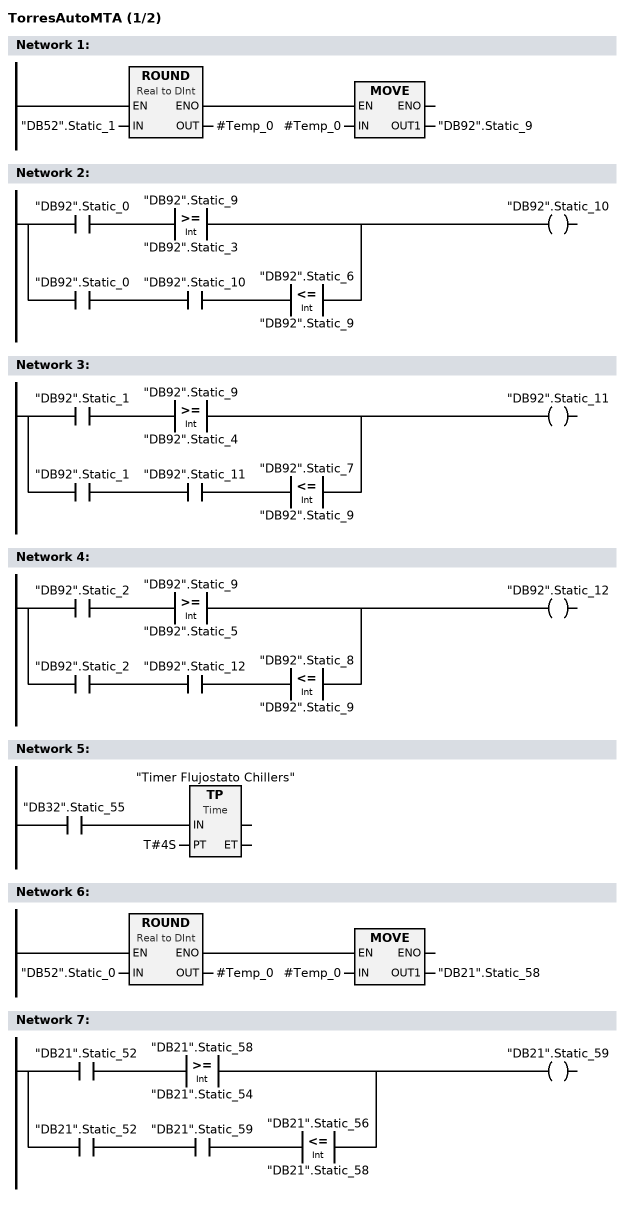
   RUNG wire#powerrail
      { S7_Templates := "[SrcType := Real, DestType := DInt]"; S7_GenerateENO := "TRUE" } Round(in := "DB52".Static_1, out => #Temp_0)
      { S7_GenerateENO := "TRUE" } Move(in := #Temp_0, out1 => "DB92".Static_9)
   END_RUNG
   // the same network as SCL:
   // ENO of a box is taken as its EN; it also drops when the box reports an error
   #Temp_0 := ROUND("DB52".Static_1);
   "DB92".Static_9 := #Temp_0;
END_REGION

REGION Network 2
   "DB92".Static_10 := ("DB92".Static_0 AND ("DB92".Static_9 >= "DB92".Static_3)) OR ("DB92".Static_0 AND "DB92".Static_10 AND ("DB92".Static_6 <= "DB92".Static_9));
END_REGION

REGION Network 3
   "DB92".Static_11 := ("DB92".Static_1 AND ("DB92".Static_9 >= "DB92".Static_4)) OR ("DB92".Static_1 AND "DB92".Static_11 AND ("DB92".Static_7 <= "DB92".Static_9));
END_REGION

REGION Network 4
   "DB92".Static_12 := ("DB92".Static_2 AND ("DB92".Static_9 >= "DB92".Static_5)) OR ("DB92".Static_2 AND "DB92".Static_12 AND ("DB92".Static_8 <= "DB92".Static_9));
END_REGION

REGION Network 5
   "Timer Flujostato Chillers".TP(pt := T#4S, in := "DB32".Static_55);
END_REGION

REGION Network 6
   RUNG wire#powerrail
      { S7_Templates := "[SrcType := Real, DestType := DInt]"; S7_GenerateENO := "TRUE" } Round(in := "DB52".Static_0, out => #Temp_0)
      { S7_GenerateENO := "TRUE" } Move(in := #Temp_0, out1 => "DB21".Static_58)
   END_RUNG
   // the same network as SCL:
   // ENO of a box is taken as its EN; it also drops when the box reports an error
   #Temp_0 := ROUND("DB52".Static_0);
   "DB21".Static_58 := #Temp_0;
END_REGION

REGION Network 7
   "DB21".Static_59 := ("DB21".Static_52 AND ("DB21".Static_58 >= "DB21".Static_54)) OR ("DB21".Static_52 AND "DB21".Static_59 AND ("DB21".Static_56 <= "DB21".Static_58));
END_REGION

REGION Network 8
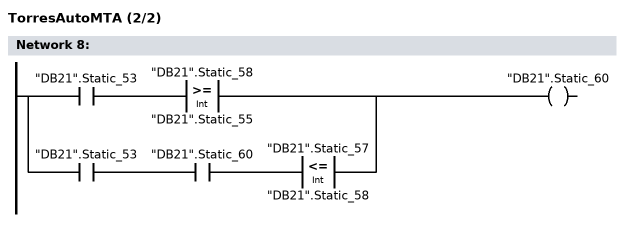
   "DB21".Static_60 := ("DB21".Static_53 AND ("DB21".Static_58 >= "DB21".Static_55)) OR ("DB21".Static_53 AND "DB21".Static_60 AND ("DB21".Static_57 <= "DB21".Static_58));
END_REGION
END_FUNCTION

(* ===== HMI "HMI_RT_3" =====
connection "Conexión2-PLC_1": ETHERNET, SIMATIC S7 300/400 MPI

HMI tags "AlarmasMTA"
   "AlarmasWord0" : Int, 1 s
   "AlarmasWord1" : Int, 1 s
   "AlarmasWord2" : Int, 1 s
   "AlarmasWord3" : Int, 1 s
   "AlarmasWord4" : Int, 1 s
   "AlarmasWord5" : Int, 1 s
   "AlarmasWord6" : Int, 1 s
   "AlarmasWord7" : Int, 1 s
   "AlarmasWord8" : Int, 1 s
   "Rec0" : Int, 1 s
   "Rec1" : Int, 1 s
   "Rec2" : Int, 1 s
   "Rec3" : Int, 1 s
   "Rec4" : Int, 1 s
   "Rec5" : Int, 1 s
   "Rec6" : Int, 1 s
   "Rec7" : Int, 1 s
   "Rec8" : Int, 1 s
   "AlarmasWord9" : Int, 1 s
   "AlarmasWord10" : Int, 1 s
   "AlarmasWord11" : Int, 1 s
   "AlarmasWord12" : Int, 1 s
   "AlarmasWord13" : Int, 1 s
   "AlarmasWord14" : Int, 1 s
   "Rec9" : Int, 1 s
   "Rec10" : Int, 1 s
   "Rec11" : Int, 1 s
   "Rec12" : Int, 1 s
   "Rec13" : Int, 1 s
   "Rec14" : Int, 1 s
   "AlarmasWord1(1)" : Int, 1 s
   "AlarmasWord15" : Int, 1 s
   "Rec15" : Int, 1 s
   "EncendidoPLC" : Bool, 1 s

HMI tags "AutoTorresChillers"
   "AutoV001" : Bool, 1 s
   "AutoV002" : Bool, 1 s
   "AutoV003" : Bool, 1 s
   "SP-ON-V001" : Int, 1 s
   "SP-ON-V002" : Int, 1 s
   "SP-ON-V003" : Int, 1 s
   "SP-OFF-V001" : Int, 1 s
   "SP-OFF-V002" : Int, 1 s
   "SP-OFF-V003" : Int, 1 s
   "TemperaturatorresCH" : Real, 1 s

HMI tags "CFG-Analog-MTA"
   "PresiónALTA" : Real, 1 s
   "PresiónBAJA" : Real, 1 s
   "TempCAV" : Real, 1 s
   "TempCH" : Real, 1 s
   "CFG-ALtaHH" : Real, 1 s
   "CFG-ALtaH" : Real, 1 s
   "CFG-ALtaL" : Real, 1 s
   "CFG-ALtaLL" : Real, 1 s
   "CFG-BajaHH" : Real, 1 s
   "CFG-BajaH" : Real, 1 s
   "CFG-BajaL" : Real, 1 s
   "CFG-BajaLL" : Real, 1 s

HMI tags "ChillersMTA"
   "HabMT007" : Bool, 1 s
   "HabMT008" : Bool, 1 s
   "HabMT009" : Bool, 1 s
   "HabMT010" : Bool, 1 s
   "DesMT007" : Bool, 1 s
   "DesMT008" : Bool, 1 s
   "DesMT009" : Bool, 1 s
   "DesMT010" : Bool, 1 s
   "MarchaMT007" : Bool, 1 s
   "MarchaMT008" : Bool, 1 s
   "MarchaMT009" : Bool, 1 s
   "MarchaMT010" : Bool, 1 s
   "ParadaMT007" : Bool, 1 s
   "ParadaMT008" : Bool, 1 s
   "ParadaMT009" : Bool, 1 s
   "ParadaMT010" : Bool, 1 s
   "Habilitación-CH-SOP-GR" : Bool, 1 s
   "Habilitación-CH-SOP-CH" : Bool, 1 s
   "Habilitación-CH-ENV-GR" : Bool, 1 s
   "Habilitación-CH-ENV-CH" : Bool, 1 s
   "Alarma1-CH-SOP-GR" : Bool, 1 s
   "Alarma2-CH-SOP-GR" : Bool, 1 s
   "RUN-CH-SOP-GR" : Bool, 1 s
   "MAX-CH-SOP-GR" : Bool, 1 s
   "AnimaciónMT007" : Byte, 1 s
   "AnimaciónMT008" : Byte, 1 s
   "AnimaciónMT009" : Byte, 1 s
   "AnimaciónMT010" : Byte, 1 s
   "AnimaciónMP010" : Byte, 1 s
   "AnimaciónMP011" : Byte, 1 s
   "AnimaciónMP012" : Byte, 1 s
   "AnimaciónMP013" : Byte, 1 s
   "HabMP010" : Bool, 1 s
   "HabMP011" : Bool, 1 s
   "HabMP012" : Bool, 1 s
   "HabMP013" : Bool, 1 s
   "HabMP018" : Bool, 1 s
   "HabMP019" : Bool, 1 s
   "DesMP010" : Bool, 1 s
   "DesMP011" : Bool, 1 s
   "DesMP012" : Bool, 1 s
   "DesMP013" : Bool, 1 s
   "DesMP018" : Bool, 1 s
   "DesMP019" : Bool, 1 s
   "MarchaMP010" : Bool, 1 s
   "MarchaMP011" : Bool, 1 s
   "MarchaMP012" : Bool, 1 s
   "MarchaMP013" : Bool, 1 s
   "MarchaMP018" : Bool, 1 s
   "MarchaMP019" : Bool, 1 s
   "ParadaMP010" : Bool, 1 s
   "ParadaMP011" : Bool, 1 s
   "ParadaMP012" : Bool, 1 s
   "ParadaMP013" : Bool, 1 s
   "ParadaMP018" : Bool, 1 s
   "ParadaMP019" : Bool, 1 s
   "AnimaciónMP018" : Byte, 1 s
   "AnimaciónMP019" : Byte, 1 s
   "DesV001" : Bool, 1 s
   "DesV002" : Bool, 1 s
   "HabV001" : Bool, 1 s
   "HabV002" : Bool, 1 s
   "MarchaV001" : Bool, 1 s
   "MarchaV002" : Bool, 1 s
   "ParadaV001" : Bool, 1 s
   "ParadaV002" : Bool, 1 s
   "AnimaciónV001" : Byte, 1 s
   "AnimaciónV002" : Byte, 1 s
   "VentiladoresMTA" : Bool, internal
   "MAX-CH-ENV-GR" : Bool, 1 s
   "RUN-CH-ENV-GR" : Bool, 1 s
   "Alarma2-CH-ENV-GR" : Bool, 1 s
   "Alarma1-CH-ENV-GR" : Bool, 1 s
   "SirenaM1" : Bool, 1 s
   "SirenaM2" : Bool, 1 s
   "SirenaM3" : Bool, 1 s
   "SirenaM4" : Bool, 1 s
   "AnimaciónV003" : Byte, 1 s
   "HabV003" : Bool, 1 s
   "DesV003" : Bool, 1 s
   "MarchaV003" : Bool, 1 s
   "ParadaV003" : Bool, 1 s
   "BombaTorreON" : Bool, 1 s
   "SirenaM5" : Bool, 1 s
   "SirenaChillers" : Bool, 1 s
   "SirenaM6" : Bool, 1 s
   "SirenaM7" : Bool, 1 s
   "SirenaM8" : Bool, 1 s
   "SirenaM9" : Bool, 1 s
   "SirenaM10" : Bool, 1 s
   "AlarmaNueva" : Bool, 1 s
   "AlarmaPresente" : Bool, 1 s
   "SinAlarmas" : Bool, 1 s
   "AlarmaAceite-CH-ENV-CH" : Bool, 1 s
   "AlarmaTemp-CH-ENV-CH" : Bool, 1 s
   "RUN-CH-ENV-CH" : Bool, 1 s
   "VerCh1MTA" : Bool, internal
   "VerCh2MTA" : Bool, internal
   "VerCh3MTA" : Bool, internal
   "VerCh4MTA" : Bool, internal
   "AlarmaPRUEBA" : DWord, 1 s
   "Presosato" : Bool, 1 s
   "CH-SOP-CH-CTC1ON" : Bool, 1 s
   "CH-SOP-CH-CTC2ON" : Bool, 1 s
   "CH-SOP-CH-TERM1" : Bool, 1 s
   "CH-SOP-CH-TERM2" : Bool, 1 s
   "CH-ENV-CH-ACT" : Bool, 1 s
   "CH-ENV-CH-TEMP" : Bool, 1 s
   "CH-ENV-CH-TERM" : Bool, 1 s
   "CH-ENV-CH-RUN" : Bool, 1 s
   "BombaTorreON2" : Bool, 1 s
   "HabV001(1)" : Bool, 1 s
   "HabV002(1)" : Bool, 1 s
   "HabV003(1)" : Bool, 1 s
   "HabV4" : Bool, 1 s
   "MarchaV001(1)" : Bool, 1 s
   "MarchaV002(1)" : Bool, 1 s
   "MarchaV003(1)" : Bool, 1 s
   "ParadaV001(1)" : Bool, 1 s
   "ParadaV002(1)" : Bool, 1 s
   "ParadaV003(1)" : Bool, 1 s
   "AnimaMenuV001" : Int, 1 s
   "AnimaMenuV002" : Int, 1 s
   "AnimaMenuV003" : Int, 1 s
   "DeshV001" : Bool, 1 s
   "DeshV002" : Bool, 1 s
   "DeshV003" : Bool, 1 s

discrete alarms
   125: '', class MTA, trigger "AlarmasWord4" bit 8
   126: '', class MTA, trigger "AlarmasWord3" bit 15
   127: '', class MTA, trigger "AlarmasWord4" bit 11
   128: '', class MTA, trigger "AlarmasWord4" bit 10
   129: '', class MTA, trigger "AlarmasWord4" bit 9
   130: '', class MTA, trigger "AlarmasWord3" bit 11
   131: '', class MTA, trigger "AlarmasWord3" bit 10
   132: '', class MTA, trigger "AlarmasWord3" bit 9
   133: '', class MTA, trigger "AlarmasWord3" bit 14
   134: '', class MTA, trigger "AlarmasWord3" bit 13
   135: '', class MTA, trigger "AlarmasWord3" bit 12
   136: '', class MTA, trigger "AlarmasWord4" bit 12
   137: '', class MTA, trigger "AlarmasWord4" bit 15
   138: '', class MTA, trigger "AlarmasWord4" bit 14
   139: '', class MTA, trigger "AlarmasWord4" bit 13
   140: '', class MTA, trigger "AlarmasWord3" bit 8
   141: '', class MTA, trigger "AlarmasWord1" bit 8
   144: '', class MTA, trigger "AlarmasWord1" bit 11
   145: '', class MTA, trigger "AlarmasWord1" bit 10
   146: '', class MTA, trigger "AlarmasWord1" bit 9
   153: '', class MTA, trigger "AlarmasWord1" bit 12
   154: '', class MTA, trigger "AlarmasWord2" bit 12
   155: '', class MTA, trigger "AlarmasWord2" bit 11
   156: '', class MTA, trigger "AlarmasWord2" bit 10
   157: '', class MTA, trigger "AlarmasWord2" bit 15
   158: '', class MTA, trigger "AlarmasWord2" bit 14
   159: '', class MTA, trigger "AlarmasWord2" bit 13
   160: '', class MTA, trigger "AlarmasWord1" bit 15
   161: '', class MTA, trigger "AlarmasWord1" bit 14
   162: '', class MTA, trigger "AlarmasWord1" bit 13
   163: '', class MTA, trigger "AlarmasWord2" bit 9
   164: '', class MTA, trigger "AlarmasWord2" bit 8
   165: '', class MTA, trigger "AlarmasWord5" bit 8
   166: '', class MTA, trigger "AlarmasWord5" bit 9
   167: '', class MTA, trigger "AlarmasWord5" bit 10
   168: '', class MTA, trigger "AlarmasWord5" bit 11
   169: '', class MTA, trigger "AlarmasWord5" bit 12
   170: '', class MTA, trigger "AlarmasWord5" bit 13
   171: '', class MTA, trigger "AlarmasWord5" bit 14
   172: '', class MTA, trigger "AlarmasWord5" bit 15
   13: '', class MTA, trigger "AlarmasWord6" bit 8
   14: '', class MTA, trigger "AlarmasWord6" bit 9
   50: '', class MTA, trigger "AlarmasWord6" bit 10
   53: '', class MTA, trigger "AlarmasWord6" bit 11
   87: '', class MTA, trigger "AlarmasWord6" bit 12
   88: '', class MTA, trigger "AlarmasWord6" bit 13
   89: '', class MTA, trigger "AlarmasWord6" bit 14
   90: '', class MTA, trigger "AlarmasWord6" bit 15
   69: '', class MTA, trigger "AlarmasWord7" bit 11
   68: '', class MTA, trigger "AlarmasWord7" bit 10
   67: '', class MTA, trigger "AlarmasWord7" bit 9
   66: '', class MTA, trigger "AlarmasWord7" bit 8
   70: '', class MTA, trigger "AlarmasWord7" bit 12
   71: '', class MTA, trigger "AlarmasWord7" bit 13
   72: '', class MTA, trigger "AlarmasWord7" bit 14
   73: '', class MTA, trigger "AlarmasWord7" bit 15
   74: '', class MTA, trigger "AlarmasWord8" bit 8
   75: '', class MTA, trigger "AlarmasWord8" bit 9
   76: '', class MTA, trigger "AlarmasWord8" bit 10
   77: '', class MTA, trigger "AlarmasWord8" bit 11
   78: '', class MTA, trigger "AlarmasWord8" bit 12
   79: '', class MTA, trigger "AlarmasWord8" bit 13
   80: '', class MTA, trigger "AlarmasWord8" bit 14
   81: '', class MTA, trigger "AlarmasWord8" bit 15
   82: '', class MTA, trigger "AlarmasWord9" bit 8
   83: '', class MTA, trigger "AlarmasWord9" bit 9
   91: '', class MTA, trigger "AlarmasWord9" bit 10
   92: '', class MTA, trigger "AlarmasWord9" bit 11
   93: '', class MTA, trigger "AlarmasWord9" bit 12
   94: '', class MTA, trigger "AlarmasWord9" bit 13
   96: '', class MTA, trigger "AlarmasWord9" bit 15
   97: '', class MTA, trigger "AlarmasWord10" bit 8
   98: '', class MTA, trigger "AlarmasWord10" bit 9
   99: '', class MTA, trigger "AlarmasWord10" bit 10
   100: '', class MTA, trigger "AlarmasWord10" bit 11
   101: '', class MTA, trigger "AlarmasWord10" bit 12
   102: '', class MTA, trigger "AlarmasWord10" bit 13
   121: '', class MTA, trigger "AlarmasWord10" bit 14
   104: '', class MTA, trigger "AlarmasWord10" bit 15
   105: '', class MTA, trigger "AlarmasWord11" bit 8
   106: '', class MTA, trigger "AlarmasWord11" bit 9
   107: '', class MTA, trigger "AlarmasWord11" bit 10
   108: '', class MTA, trigger "AlarmasWord11" bit 11
   109: '', class MTA, trigger "AlarmasWord11" bit 12
   110: '', class MTA, trigger "AlarmasWord11" bit 13
   111: '', class MTA, trigger "AlarmasWord11" bit 14
   112: '', class MTA, trigger "AlarmasWord11" bit 15
   113: '', class MTA, trigger "AlarmasWord12" bit 8
   114: '', class MTA, trigger "AlarmasWord12" bit 9
   115: '', class MTA, trigger "AlarmasWord12" bit 10
   116: '', class MTA, trigger "AlarmasWord12" bit 11
   117: '', class MTA, trigger "AlarmasWord12" bit 12
   118: '', class MTA, trigger "AlarmasWord12" bit 13
   119: '', class MTA, trigger "AlarmasWord12" bit 14
   120: '', class MTA, trigger "AlarmasWord12" bit 15
   122: '', class MTA, trigger "AlarmasWord13" bit 8
   1: '', class MTA, trigger "AlarmasWord13" bit 9
   2: '', class MTA, trigger "AlarmasWord13" bit 10
   3: '', class MTA, trigger "AlarmasWord13" bit 11
   4: '', class MTA, trigger "AlarmasWord13" bit 12
   5: '', class MTA, trigger "AlarmasWord13" bit 13
   6: '', class MTA, trigger "AlarmasWord13" bit 14
   7: '', class MTA, trigger "AlarmasWord13" bit 15
   8: '', class MTA, trigger "AlarmasWord14" bit 8
   9: '', class MTA, trigger "AlarmasWord14" bit 9
   10: '', class MTA, trigger "AlarmasWord14" bit 10
   11: '', class MTA, trigger "AlarmasWord14" bit 11
   12: '', class MTA, trigger "AlarmasWord14" bit 12
   15: '', class MTA, trigger "AlarmasWord14" bit 13
   16: '', class MTA, trigger "AlarmasWord14" bit 14
   17: '', class MTA, trigger "AlarmasWord14" bit 15
   95: '', class MTA, trigger "AlarmasWord9" bit 14
   149: '', class MTA, trigger "AlarmasWord0" bit 8
   142: '', class MTA, trigger "AlarmasWord0" bit 15
   143: '', class MTA, trigger "AlarmasWord0" bit 14
   152: '', class MTA, trigger "AlarmasWord0" bit 11
   147: '', class MTA, trigger "AlarmasWord0" bit 10
   148: '', class MTA, trigger "AlarmasWord0" bit 9
   150: '', class MTA, trigger "AlarmasWord0" bit 13
   151: '', class MTA, trigger "AlarmasWord0" bit 12
   21: '', class MTA, trigger "AlarmasWord15" bit 11
   22: '', class MTA, trigger "AlarmasWord15" bit 12
   19: '', class MTA, trigger "AlarmasWord15" bit 9
   20: '', class MTA, trigger "AlarmasWord15" bit 10
   23: '', class MTA, trigger "AlarmasWord15" bit 13
   24: '', class MTA, trigger "AlarmasWord15" bit 14
   25: '', class MTA, trigger "AlarmasWord15" bit 15
   18: '', class MTA, trigger "AlarmasWord15" bit 8

text list "EstadoMotor": 0 ''; 1 ''; 2 ''; 3 ''; 4 ''; 5 ''; 6 ''; 7 ''

graphic list "Motor2": 0 'Motor2Dorado'; 1 'Motor2Verde_1'; 2 'Motor2VerdeOscuro'; 3 'Motor2Azul'; 4 'Motor2Celeste'; 5 'Motor2Amarillo'; 6 'Motor2Gris_1'; 7 'Motor2Rojo'

graphic list "MotorTorre": 0 'torreFINAL4C2_1'; 1 'torreFINAL4C2v_2'; 2 'torreFINAL4C2v_2'; 3 'torreFINAL4C2b'; 4 'torreFINAL4C2b'; 5 'torreFINAL4C2a_2'; 6 'torreFINAL4C2_1'; 7 'torreFINAL4C2_1'

graphic list "Indicador": 0 'indDorado'; 1 'indVerde'; 2 'indVerde_1'; 3 'indAZUL'; 4 'indCeleste'; 5 'indAmarillo'; 6 'indGris'; 7 'indRojo'

graphic list "Secador2": 0 'BaseSullChicoDorado_2'; 1 'BaseSullChico_5'; 2 'BaseSullChico_5'; 3 'BaseSullChicoAzul_2'; 4 'BaseSullChicoAzul_2'; 5 'BaseSullChicoAmarillo_2'; 6 'BaseSullChicoGris_2'; 7 'BaseSullChicoRojo_2'

graphic list "Secador3": 0 'BaseSullChicoDorado_3'; 1 'BaseSullChico_6'; 2 'BaseSullChico_6'; 3 'BaseSullChicoAzul_3'; 4 'BaseSullChicoAzul_3'; 5 'BaseSullChicoAmarillo_3'; 6 'BaseSullChicoGris_3'; 7 'BaseSullChicoRojo_3'

graphic list "Secador1": 0 'BaseSullChicoDorado_1'; 1 'BaseSullChico_4'; 2 'BaseSullChico_4'; 3 'BaseSullChicoAzul_1'; 4 'BaseSullChicoAzul_1'; 5 'BaseSullChicoAmarillo_1'; 6 'BaseSullChicoGris_1'; 7 'BaseSullChicoRojo_1'

screen "MTA-Avisos" 800x480, template "Plantilla_2"
   AlarmView "Visor de avisos_1" at 5,53 size 790x367
   TextField "Campo de texto_5" at 327,10 size 54x27

screen "MTA-ChillersBombasEnvasado" 800x480, template "Plantilla_2"
   GraphicView "Visor de gráficos_3" at 648,158 size 48x71
   GraphicIOField "Plantilla_Campo ES gráfico_2" at 684,217 size 49x36
   SymbolicIOField "Campo ES simbólico_4" at 602,132 size 172x21
   TextField "Campo de texto_6" at 599,93 size 42x18
   GraphicView "Visor de gráficos_4" at 454,158 size 48x71
   GraphicIOField "Plantilla_Campo ES gráfico_1" at 490,217 size 49x36
   SymbolicIOField "Campo ES simbólico_1" at 408,132 size 172x21
   TextField "Campo de texto_7" at 405,93 size 42x18
   GraphicView "Visor de gráficos_6" at 64,158 size 48x71
   GraphicIOField "Plantilla_Campo ES gráfico_4" at 100,217 size 49x36
   SymbolicIOField "Campo ES simbólico_3" at 20,132 size 172x21
   TextField "Campo de texto_9" at 23,93 size 41x18
   TextField "Campo de texto_19" at 405,112 size 169x18
   GraphicView "Visor de gráficos_5" at 260,158 size 48x71
   GraphicIOField "Plantilla_Campo ES gráfico_3" at 296,217 size 49x36
   SymbolicIOField "Campo ES simbólico_2" at 214,132 size 172x21
   TextField "Campo de texto_8" at 211,93 size 41x18
   TextField "Campo de texto_18" at 598,112 size 150x18
   TextField "Campo de texto_16" at 215,113 size 150x18
   TextField "Campo de texto_17" at 21,113 size 146x18
   GraphicView "Plantilla_Visor de gráficos_2" at 752,6 size 35x35
   GraphicView "Plantilla_Visor de gráficos_1" at 752,6 size 35x35
   Button "Botón_1" at 740,1 size 57x44
   ScreenModuleView "ControlMotor-NoAUTO_1" at 609,271 size 163x76
   ScreenModuleView "ControlMotor-NoAUTO_2" at 413,271 size 163x76
   ScreenModuleView "ControlMotor-NoAUTO_3" at 219,271 size 163x76
   ScreenModuleView "ControlMotor-NoAUTO_4" at 22,271 size 163x76
   TextField "Campo de texto_5" at 256,10 size 261x27

screen "MTA-ChillersBombasSoplado" 800x480, template "Plantilla_2"
   TextField "Campo de texto_5" at 256,10 size 248x27
   GraphicView "Visor de gráficos_3" at 648,158 size 48x71
   GraphicIOField "Plantilla_Campo ES gráfico_8" at 684,217 size 49x36
   SymbolicIOField "Campo ES simbólico_4" at 602,132 size 172x21
   TextField "Campo de texto_6" at 599,93 size 42x18
   GraphicView "Visor de gráficos_4" at 454,158 size 48x71
   GraphicIOField "Plantilla_Campo ES gráfico_7" at 490,217 size 49x36
   SymbolicIOField "Campo ES simbólico_1" at 408,132 size 172x21
   TextField "Campo de texto_7" at 405,93 size 42x18
   GraphicView "Visor de gráficos_6" at 64,158 size 48x71
   GraphicIOField "Plantilla_Campo ES gráfico_5" at 100,217 size 49x36
   SymbolicIOField "Campo ES simbólico_3" at 20,132 size 172x21
   TextField "Campo de texto_9" at 23,93 size 41x18
   TextField "Campo de texto_19" at 407,113 size 140x18
   GraphicView "Visor de gráficos_5" at 260,158 size 48x71
   GraphicIOField "Plantilla_Campo ES gráfico_6" at 296,217 size 49x36
   SymbolicIOField "Campo ES simbólico_2" at 214,132 size 172x21
   TextField "Campo de texto_8" at 211,93 size 41x18
   TextField "Campo de texto_18" at 599,113 size 104x18
   TextField "Campo de texto_16" at 212,113 size 142x18
   TextField "Campo de texto_17" at 21,113 size 138x18
   GraphicView "Plantilla_Visor de gráficos_2" at 752,6 size 35x35
   GraphicView "Plantilla_Visor de gráficos_1" at 752,6 size 35x35
   Button "Botón_1" at 740,1 size 57x44
   ScreenModuleView "ControlMotor-NoAUTO_1" at 609,271 size 163x76
   ScreenModuleView "ControlMotor-NoAUTO_3" at 219,271 size 163x76
   ScreenModuleView "ControlMotor-NoAUTO_2" at 417,271 size 163x76
   ScreenModuleView "ControlMotor-NoAUTO_4" at 27,271 size 163x76

screen "MTA-ChillersConfiguraciónSirena" 800x480, template "Plantilla_2"
   Switch "Interruptor_1" at 119,81 size 36x32
   Switch "Interruptor_2" at 119,118 size 36x32
   Switch "Interruptor_3" at 119,155 size 36x32
   Switch "Interruptor_4" at 119,192 size 36x32
   Switch "Interruptor_5" at 119,229 size 36x32
   TextField "Campo de texto_1" at 163,233 size 365x22
   TextField "Campo de texto_2" at 163,196 size 424x22
   TextField "Campo de texto_3" at 163,160 size 353x22
   TextField "Campo de texto_4" at 163,122 size 411x22
   TextField "Campo de texto_5" at 163,86 size 340x22
   TextField "Campo de texto_6" at 51,53 size 277x22
   TextField "Campo de texto_7" at 214,8 size 319x29
   Switch "Interruptor_6" at 119,266 size 36x32
   TextField "Campo de texto_8" at 163,271 size 231x22
   Switch "Interruptor_7" at 119,303 size 36x32
   TextField "Campo de texto_9" at 163,307 size 244x22
   Switch "Interruptor_8" at 119,341 size 36x32
   TextField "Campo de texto_10" at 163,346 size 150x22
   GraphicView "Plantilla_Visor de gráficos_2" at 752,6 size 35x35
   GraphicView "Plantilla_Visor de gráficos_1" at 752,6 size 35x35
   Button "Botón_1" at 740,1 size 57x44
   Switch "Interruptor_9" at 119,378 size 36x32
   TextField "Campo de texto_11" at 163,383 size 194x22

screen "MTA-Chillers-Envasado" 800x480, template "Plantilla_2"
   GraphicView "Visor de gráficos_2" at 24,127 size 192x232
   GraphicView "Visor de gráficos_1" at 432,129 size 144x104
   Switch "Interruptor_1" at 243,127 size 91x31
   TextField "Campo de texto_5" at 309,10 size 182x27
   TextField "Campo de texto_10" at 19,78 size 169x22
   TextField "Campo de texto_6" at 411,78 size 158x22
   TextField "Campo de texto_1" at 263,203 size 40x18
   TextField "Campo de texto_3" at 263,182 size 108x18
   TextField "Campo de texto_4" at 263,223 size 101x18
   Switch "Interruptor_2" at 595,127 size 91x31
   GraphicView "Plantilla_Visor de gráficos_2" at 752,6 size 35x35
   GraphicView "Plantilla_Visor de gráficos_1" at 752,6 size 35x35
   Button "Botón_1" at 740,1 size 57x44
   TextField "Campo de texto_24" at 613,183 size 79x18
   TextField "Campo de texto_25" at 613,166 size 108x18
   TextField "Campo de texto_26" at 613,201 size 115x18
   TextField "Campo de texto_27" at 613,220 size 125x18

screen "MTA-Chillers-General" 800x480, template "Plantilla_2"
   GraphicView "Visor de gráficos_7" at 488,183 size 48x71
   GraphicView "Visor de gráficos_8" at 536,183 size 48x71
   GraphicView "Visor de gráficos_1" at 392,183 size 48x71
   GraphicView "Visor de gráficos_9" at 440,183 size 48x71
   GraphicView "Visor de gráficos_17" at 383,130 size 87x77
   GraphicView "Visor de gráficos_18" at 479,130 size 87x77
   GraphicView "Visor de gráficos_14" at 384,48 size 141x131
   GraphicView "Visor de gráficos_3" at 750,189 size 48x212
   GraphicView "Visor de gráficos_4" at 630,161 size 96x96
   GraphicView "Visor de gráficos_5" at 264,183 size 48x71
   GraphicView "Visor de gráficos_6" at 312,183 size 48x71
   GraphicView "Visor de gráficos_10" at 168,183 size 48x71
   GraphicView "Visor de gráficos_11" at 216,183 size 48x71
   GraphicView "Visor de gráficos_2" at 12,132 size 128x144
   GraphicView "Visor de gráficos_12" at 45,333 size 88x77
   GraphicView "Visor de gráficos_15" at 159,130 size 87x77
   GraphicView "Visor de gráficos_16" at 255,130 size 87x77
   GraphicView "Visor de gráficos_13" at 162,48 size 141x131
   GraphicIOField "Plantilla_Campo ES gráfico_2" at 304,240 size 41x36
   GraphicIOField "Plantilla_Campo ES gráfico_1" at 352,240 size 41x36
   GraphicIOField "Plantilla_Campo ES gráfico_3" at 528,240 size 41x36
   GraphicIOField "Plantilla_Campo ES gráfico_4" at 576,240 size 41x36
   GraphicIOField "Plantilla_Campo ES gráfico_5" at 432,240 size 41x36
   GraphicIOField "Plantilla_Campo ES gráfico_6" at 480,240 size 41x36
   GraphicIOField "Plantilla_Campo ES gráfico_7" at 208,240 size 41x36
   GraphicIOField "Plantilla_Campo ES gráfico_8" at 256,240 size 41x36
   TextField "Campo de texto_1" at 631,124 size 86x32
   TextField "Campo de texto_2" at 668,364 size 86x32
   TextField "Campo de texto_3" at 142,373 size 90x32
   TextField "Campo de texto_4" at 28,94 size 90x32
   TextField "Campo de texto_5" at 334,8 size 72x29
   TextField "Campo de texto_6" at 474,309 size 131x25
   TextField "Campo de texto_7" at 242,309 size 139x25
   TextField "Campo de texto_9" at 520,70 size 51x52
   TextField "Campo de texto_8" at 214,277 size 41x19
   TextField "Campo de texto_11" at 262,277 size 41x19
   TextField "Campo de texto_12" at 310,277 size 49x19
   TextField "Campo de texto_13" at 366,277 size 42x19
   TextField "Campo de texto_14" at 438,277 size 41x19
   TextField "Campo de texto_15" at 486,277 size 41x19
   TextField "Campo de texto_16" at 534,277 size 42x19
   TextField "Campo de texto_17" at 590,277 size 42x19
   TextField "Campo de texto_10" at 294,69 size 58x52
   Button "Botón_3" at 629,155 size 170x254
   Button "Botón_2" at 419,227 size 215x78
   Button "Botón_4" at 0,122 size 194x294
   Button "Botón_5" at 203,226 size 208x79
   GraphicView "Plantilla_Visor de gráficos_2" at 752,6 size 35x35
   GraphicView "Plantilla_Visor de gráficos_1" at 752,6 size 35x35
   Button "Botón_1" at 740,1 size 57x44

screen "MTA-Chillers-Soplado" 800x480, template "Plantilla_2"
   GraphicView "Visor de gráficos_2" at 24,127 size 192x232
   GraphicView "Visor de gráficos_1" at 424,129 size 160x168
   Switch "Interruptor_1" at 243,127 size 91x31
   TextField "Campo de texto_1" at 263,203 size 40x18
   TextField "Campo de texto_3" at 263,182 size 108x18
   TextField "Campo de texto_4" at 263,223 size 101x18
   TextField "Campo de texto_5" at 311,10 size 169x27
   TextField "Campo de texto_10" at 19,78 size 156x22
   TextField "Campo de texto_6" at 411,78 size 145x22
   Switch "Interruptor_2" at 627,127 size 91x31
   GraphicView "Plantilla_Visor de gráficos_2" at 752,6 size 35x35
   GraphicView "Plantilla_Visor de gráficos_1" at 752,6 size 35x35
   Button "Botón_1" at 740,1 size 57x44
   TextField "Campo de texto_28" at 607,198 size 120x18
   TextField "Campo de texto_29" at 607,177 size 120x18
   TextField "Campo de texto_30" at 631,220 size 96x18
   TextField "Campo de texto_31" at 631,241 size 96x18

screen "MTA-TorreEnfriamientoBMB" 800x480, template "Plantilla_2"
   GraphicView "Visor de gráficos_1" at 167,153 size 98x119
   GraphicView "Visor de gráficos_4" at 260,143 size 138x153
   GraphicView "Visor de gráficos_17" at 16,128 size 178x201
   GraphicView "Visor de gráficos_2" at 167,153 size 98x119
   GraphicView "Visor de gráficos_3" at 260,143 size 138x153
   GraphicView "Visor de gráficos_5" at 16,128 size 178x201
   GraphicView "Visor de gráficos_6" at 167,153 size 98x119
   GraphicView "Visor de gráficos_15" at 260,143 size 138x153
   GraphicView "Visor de gráficos_16" at 16,128 size 178x201
   TextField "Campo de texto_1" at 361,84 size 57x23
   TextField "Campo de texto_2" at 229,95 size 47x20
   TextField "Campo de texto_12" at 101,76 size 57x23
   TextField "Campo de texto_13" at 273,197 size 55x29
   TextField "Campo de texto_14" at 38,202 size 50x34
   GraphicIOField "Campo ES gráfico_1" at 76,122 size 56x29
   GraphicIOField "Campo ES gráfico_2" at 199,147 size 33x21
   GraphicIOField "Campo ES gráfico_3" at 306,137 size 45x24
   GraphicView "Visor de gráficos_19" at 0,384 size 800x15
   GraphicView "Plantilla_Visor de gráficos_2" at 752,6 size 35x35
   GraphicView "Plantilla_Visor de gráficos_1" at 752,6 size 35x35
   Button "Botón_1" at 740,1 size 57x44
   Button "Botón_2" at 200,320 size 152x38
   TextField "Campo de texto_10" at 41,374 size 98x32
   TextField "Campo de texto_5" at 238,8 size 293x29
   GraphicView "Visor de gráficos_9" at 30,56 size 63x62
   GraphicView "Visor de gráficos_10" at 30,56 size 63x62
   GraphicView "Visor de gráficos_11" at 177,82 size 47x46
   GraphicView "Visor de gráficos_12" at 177,82 size 47x46
   GraphicView "Visor de gráficos_13" at 292,66 size 63x62
   GraphicView "Visor de gráficos_14" at 292,66 size 63x62
   IOField "Campo ES_1" at 241,360 size 80x23
   GraphicView "Visor de gráficos_8" at 459,277 size 48x71
   GraphicIOField "Plantilla_Campo ES gráfico_1" at 497,336 size 49x36
   SymbolicIOField "Campo ES simbólico_1" at 581,259 size 172x20
   TextField "Campo de texto_7" at 495,293 size 41x18
   TextField "Campo de texto_17" at 455,241 size 129x27
   ScreenModuleView "ControlMotor-NoAUTO_4" at 565,285 size 203x76
   ScreenModuleView "ControlMotor-NoAUTO_1" at 564,115 size 203x76
   SymbolicIOField "Campo ES simbólico_4" at 575,89 size 172x20
   TextField "Campo de texto_6" at 494,129 size 41x18
   TextField "Campo de texto_16" at 454,77 size 151x27
   GraphicView "Visor de gráficos_7" at 458,113 size 48x71
   GraphicIOField "Plantilla_Campo ES gráfico_2" at 496,172 size 49x36

screen "MTA-TorreEnfriamientoVENT" 800x480, template "Plantilla_2"
   GraphicView "Visor de gráficos_1" at 167,153 size 98x119
   GraphicView "Visor de gráficos_4" at 260,143 size 138x153
   GraphicView "Visor de gráficos_17" at 16,128 size 178x201
   GraphicView "Visor de gráficos_2" at 167,153 size 98x119
   GraphicView "Visor de gráficos_3" at 260,143 size 138x153
   GraphicView "Visor de gráficos_5" at 16,128 size 178x201
   GraphicView "Visor de gráficos_6" at 167,153 size 98x119
   GraphicView "Visor de gráficos_15" at 260,143 size 138x153
   GraphicView "Visor de gráficos_16" at 16,128 size 178x201
   SymbolicIOField "Campo ES simbólico_2" at 548,59 size 188x19
   SymbolicIOField "Campo ES simbólico_3" at 549,181 size 188x19
   SymbolicIOField "Campo ES simbólico_7" at 549,301 size 188x19
   TextField "Campo de texto_1" at 361,84 size 57x23
   TextField "Campo de texto_2" at 229,95 size 47x20
   TextField "Campo de texto_13" at 273,197 size 55x29
   TextField "Campo de texto_14" at 38,202 size 50x34
   ScreenModuleView "Faceplate_4_1" at 447,84 size 245x68
   TextField "Campo de texto_4" at 439,176 size 104x27
   TextField "Campo de texto_3" at 439,54 size 104x27
   TextField "Campo de texto_23" at 440,298 size 104x27
   ScreenModuleView "Faceplate_4_2" at 447,204 size 245x68
   ScreenModuleView "Faceplate_4_3" at 447,326 size 245x68
   TextField "Campo de texto_12" at 101,76 size 57x23
   GraphicIOField "Campo ES gráfico_1" at 76,122 size 56x29
   GraphicIOField "Campo ES gráfico_2" at 199,147 size 33x21
   GraphicIOField "Campo ES gráfico_3" at 306,137 size 45x24
   Switch "Interruptor_1" at 744,62 size 32x29
   Switch "Interruptor_2" at 744,184 size 32x29
   Switch "Interruptor_3" at 744,304 size 32x29
   GraphicView "Visor de gráficos_19" at 0,384 size 800x15
   TextField "Campo de texto_5" at 238,8 size 293x29
   GraphicView "Visor de gráficos_9" at 30,56 size 63x62
   GraphicView "Visor de gráficos_10" at 30,56 size 63x62
   GraphicView "Visor de gráficos_11" at 177,82 size 47x46
   GraphicView "Visor de gráficos_12" at 177,82 size 47x46
   GraphicView "Visor de gráficos_13" at 292,66 size 63x62
   GraphicView "Visor de gráficos_14" at 292,66 size 63x62
   GraphicView "Plantilla_Visor de gráficos_2" at 752,6 size 35x35
   GraphicView "Plantilla_Visor de gráficos_1" at 752,6 size 35x35
   Button "Botón_1" at 740,1 size 57x44
   TextField "Campo de texto_10" at 41,374 size 98x32
   Button "Botón_2" at 200,320 size 152x38
   IOField "Campo ES_1" at 241,360 size 80x23
   GraphicIOField "Campo ES gráfico_4" at 429,160 size 362x6
   GraphicIOField "Campo ES gráfico_5" at 429,282 size 362x6
   GraphicIOField "Campo ES gráfico_6" at 429,404 size 362x6

Template "Plantilla_2" 800x480
   Button "Plantilla_1" at 640,429 size 78x48
   Button "Plantilla_8" at 81,429 size 78x48
   Button "Plantilla_10" at 2,429 size 78x48
   Button "Plantilla_11" at 720,429 size 78x48
   Button "Plantilla_2" at 480,429 size 78x48
   Button "Plantilla_3" at 560,429 size 78x48
   Button "Plantilla_4" at 400,429 size 78x48
   Button "Plantilla_5" at 320,429 size 78x48
   Button "Plantilla_6" at 240,429 size 78x48
   Button "Plantilla_7" at 160,429 size 78x48
   GraphicView "Plantilla_Visor de gráficos_26" at 68,9 size 91x26
   GraphicView "Plantilla_Visor de gráficos_27" at 9,8 size 49x29
*)

(* ===== HMI "HMI_RT_1" =====

text list "Enclavamientos": 0 ''; 1 ''; 2 ''; 3 ''; 4 ''; 5 ''

ScreenModuleEditorView "Faceplate_7" 640x480
   GraphicView "Visor de gráficos_1" at 10,10 size 143x70
   GraphicView "Visor de gráficos_2" at 10,10 size 143x70
*)

(* ===== HMI "HMI_RT_1" =====

text list "EstadoMotor": 0 ''; 1 ''; 2 ''; 3 ''; 4 ''; 5 ''; 6 ''; 7 ''